FUNCTION_BLOCK PreemptivePriority
VAR_INPUT
  xCondition : ARRAY [1..13] OF BOOL;  (* 条件1 *)
  xTaskComplete : BOOL;  (* 任务完成 *)
  xReset : BOOL;  (* 复位 *)
END_VAR
VAR
  xOccupy : BOOL;  (* 占用 *)
END_VAR
VAR_OUTPUT
  iPriority : INT;  (* 输出任务号 *)
END_VAR
VAR
  m_tonConditionDelay : TON;
  m_xConditionDelay : BOOL;
  m_tConditionCurrentTime : TIME;
  m_iLastTask : INT;  (* 上次执行的任务 *)
  m_tpLastTaskPulse1 : TP;
  m_tpLastTaskPulse2 : TP;
  m_tpLastTaskPulse3 : TP;
  m_tpLastTaskPulse4 : TP;
  m_tpLastTaskPulse5 : TP;
  m_xLastTaskPulse : ARRAY [1..13] OF BOOL;
  m_tLastTaskPulse : ARRAY [1..13] OF TIME := [13(T#0s)];
  m_tpLastTaskPulse6 : TON;
  ii : INT;
END_VAR
VAR CONSTANT
  CONDITION_QUANTITY : INT := 13;
END_VAR
VAR
  m_tpLastTaskPulse7 : TON;
  m_tpLastTaskPulse8 : TON;
  m_tpLastTaskPulse9 : TON;
  m_tpLastTaskPulse10 : TON;
  m_tpLastTaskPulse11 : TON;
  m_tpLastTaskPulse12 : TON;
  m_tpLastTaskPulse13 : TON;
END_VAR
(*抢占式优先级块
现在满足13个条件的任务进行抢占式优先级排列
条件满足后延时两秒，开始执行任务，
同一任务连续执行优先级下降
需要改造成任意多个
使用于一个入口多个出口的程序，使用抢占式优先级块
*)
IF LDP(TRUE, xTaskComplete) THEN
	xOccupy:=0;
	iPriority:=0;
END_IF;
(*//任务滤波，延时两秒*)
m_tonConditionDelay(IN:=( xCondition[1]
						OR xCondition[2]
						OR xCondition[3]
						OR xCondition[4]
						OR xCondition[5]
						OR xCondition[6]
						OR xCondition[7]
						OR xCondition[8]
						OR xCondition[9]
						OR xCondition[10]
						OR xCondition[11]
						OR xCondition[12]
						OR xCondition[13]
						)
						AND iPriority=0,
					PT:= T#1s,
					Q:= m_xConditionDelay ,
					ET:= m_tConditionCurrentTime );		
(*//判断优先级，上个任务与本次任务相同，延时一秒执行*)
m_tpLastTaskPulse1(IN:= xCondition[1]  AND m_iLastTask=1 AND m_xConditionDelay  ,PT:= T#1s,Q:= m_xLastTaskPulse[1],ET:= m_tLastTaskPulse[1] );
m_tpLastTaskPulse2(IN:= xCondition[2]  AND m_iLastTask=2 AND m_xConditionDelay  ,PT:= T#1s,Q:= m_xLastTaskPulse[2],ET:= m_tLastTaskPulse[2] );
m_tpLastTaskPulse3(IN:= xCondition[3]  AND m_iLastTask=3 AND m_xConditionDelay  ,PT:= T#1s,Q:= m_xLastTaskPulse[3],ET:= m_tLastTaskPulse[3] );
m_tpLastTaskPulse4(IN:= xCondition[4]  AND m_iLastTask=4 AND m_xConditionDelay  ,PT:= T#1s,Q:= m_xLastTaskPulse[4],ET:= m_tLastTaskPulse[4] );
m_tpLastTaskPulse5(IN:= xCondition[5]  AND m_iLastTask=5 AND m_xConditionDelay  ,PT:= T#1s,Q:= m_xLastTaskPulse[5],ET:= m_tLastTaskPulse[5] );
m_tpLastTaskPulse6(IN:= xCondition[6]  AND m_iLastTask=6 AND m_xConditionDelay  ,PT:= T#1s,Q:= m_xLastTaskPulse[6],ET:= m_tLastTaskPulse[6] );
m_tpLastTaskPulse7(IN:= xCondition[7]  AND m_iLastTask=7 AND m_xConditionDelay  ,PT:= T#1s,Q:= m_xLastTaskPulse[7],ET:= m_tLastTaskPulse[7] );
m_tpLastTaskPulse8(IN:= xCondition[8]  AND m_iLastTask=8 AND m_xConditionDelay  ,PT:= T#1s,Q:= m_xLastTaskPulse[8],ET:= m_tLastTaskPulse[8] );
m_tpLastTaskPulse9(IN:= xCondition[9]  AND m_iLastTask=9 AND m_xConditionDelay  ,PT:= T#1s,Q:= m_xLastTaskPulse[9],ET:= m_tLastTaskPulse[9] );
m_tpLastTaskPulse10(IN:= xCondition[10]  AND m_iLastTask=10 AND m_xConditionDelay  ,PT:= T#1s,Q:= m_xLastTaskPulse[10],ET:= m_tLastTaskPulse[10] );
m_tpLastTaskPulse11(IN:= xCondition[11]  AND m_iLastTask=11 AND m_xConditionDelay  ,PT:= T#1s,Q:= m_xLastTaskPulse[11],ET:= m_tLastTaskPulse[11] );
m_tpLastTaskPulse12(IN:= xCondition[12]  AND m_iLastTask=12 AND m_xConditionDelay  ,PT:= T#1s,Q:= m_xLastTaskPulse[12],ET:= m_tLastTaskPulse[12] );
m_tpLastTaskPulse13(IN:= xCondition[13]  AND m_iLastTask=13 AND m_xConditionDelay  ,PT:= T#1s,Q:= m_xLastTaskPulse[13],ET:= m_tLastTaskPulse[13] );
(*//执行*)
FOR ii:=1 TO CONDITION_QUANTITY BY 1 DO 
	IF NOT xCondition[ii] AND NOT xOccupy THEN
		iPriority:=0;
	END_IF;
	IF xCondition[ii] AND NOT xOccupy AND m_xConditionDelay AND NOT  m_xLastTaskPulse[ii]  THEN
		iPriority:=ii;
		xOccupy:=1;
		m_iLastTask:=ii;
	END_IF;
END_FOR;        
(*//复位*)
IF xReset THEN
	iPriority:=0;
	xOccupy:=0;
	m_iLastTask:=0;	
END_IF;
(*//清除占用*)
IF iPriority=0 THEN
	xOccupy:=0;
END_IF;
END_FUNCTION_BLOCK

FUNCTION_BLOCK PriorityQueue
VAR_INPUT
  arrxCondition : ARRAY [1..13] OF QueueElement;
  xTaskComplete : BOOL;  (* 任务完成 *)
  xReset : BOOL;  (* 复位 *)
END_VAR
VAR
  xOccupy : BOOL;  (* 占用 *)
END_VAR
VAR_OUTPUT
  iPriority : INT;  (* 输出任务号 *)
END_VAR
VAR
  jj : INT;
END_VAR
VAR CONSTANT
  CONDITION_QUANTITY : INT := 3;
END_VAR
VAR
  arriTaskStack : ARRAY [0..13] OF INT;
  ii : INT;
  kk : INT;
  arrxConditionDelay : ARRAY [1..13] OF BOOL;
  arrxConditionEdgeDetect : ARRAY [1..13] OF BOOL;
  arrxDelayEdgeDetect : ARRAY [1..13] OF BOOL;
  arriDelayCounter : ARRAY [1..13] OF INT;
  ll : INT;
  Temp : INT;
  mm : INT;
  nn : INT;
  Temp2 : INT;
  oo : INT;
END_VAR
(****************************************************************************)
(*
一般情况多对一的任务调度采用这个结构，排队通过出口
优先级功能块，存储任意条件的优先级，实现栈功能先入先出，
复位功能还有问题，
出入栈式优先级块，满足条件后入栈，先入先出，在栈尾加载新任务
栈首为当前执行的任务，任务完成使用上升沿触发，触发后栈首元素弹出

复位功能清空堆栈，栈的容量在CONDITION_QUANTITY 设置
增加了结构体，结构体中带有一个条件函数，和一个优先级指示
任务完成后通过凭借优先级来排序，优先级高的条件先执行   优先级排序是从小到大的，数值小的优先级高
防止干扰，增加了任务的1秒的延时
*)

(***************************************************************************)
(*(//入栈*)
FOR ii:=1 TO CONDITION_QUANTITY BY 1 DO
	(*//循环内无法用定时器，改用计数器的形式*)
	IF arrxCondition[ii].xCondition AND SM411 (*//0.2秒的方波信号，如果移植需要修改成两个定时器*)
		AND arriDelayCounter[ii]<6  (* //计数为6，5个0.2秒的方波，所以为1秒*)
		AND NOT arrxDelayEdgeDetect[ii] THEN    (*//循环内无法用沿函数，增加锁定标志位*)
		arriDelayCounter[ii]:=arriDelayCounter[ii]+1;   (*//计数*)
	END_IF;
	IF NOT arrxCondition[ii].xCondition THEN
		arriDelayCounter[ii]:=0;   (*//计数清零*)
	END_IF;
	arrxDelayEdgeDetect[ii]:=arrxCondition[ii].xCondition AND SM411;  (*//沿函数锁，保证每次SM411为1时只记一次数*)
	IF arriDelayCounter[ii]=5 AND NOT arrxConditionEdgeDetect[ii] THEN;  (*//条件满足1秒后*)
		FOR kk:=0 TO CONDITION_QUANTITY BY 1 DO    
			IF arriTaskStack[kk]=0 THEN
				arriTaskStack[kk]:=ii;   (*//栈尾添加*)
				EXIT;
			END_IF;		
		END_FOR;
	END_IF;	
	arrxConditionEdgeDetect[ii]:=arriDelayCounter[ii]=5;  (*//边沿，这个保证只在=5时，栈尾添加一次*)
END_FOR;
(*//栈顶任务为当前执行的任务**)
iPriority:=arriTaskStack[0]; 
(*//栈顶任务完成，弹出*)
IF 	LDP(TRUE, xTaskComplete) THEN
	FOR jj:=0 TO CONDITION_QUANTITY-1 BY 1 DO
		arriTaskStack[jj]:=arriTaskStack[jj+1];
	END_FOR;
	arriTaskStack[CONDITION_QUANTITY]:=0;(*//栈尾清零*)
	(*//排序，使用插入排序*)
	FOR oo:=0 TO CONDITION_QUANTITY BY 1 DO
		IF arriTaskStack[oo]=0 THEN
			EXIT;  (* //寻找栈中不为零的元素  ，防止0元素进入条件查找的时候报错*)
		END_IF;
	END_FOR;
	(*//插入排序insertionsort*)
	FOR mm:=1 TO oo-1  BY 1 DO   (*//从1开始*)
		Temp:=arriTaskStack[mm];  (*//当前数据记录 *)
		Temp2:=arrxCondition[arriTaskStack[mm]].iPriority;  (*//当前优先级记录 *)
		nn:=mm;  (*//指针赋值*)
		WHILE  (nn>0 AND Temp2< arrxCondition[arriTaskStack[nn-1]].iPriority)  DO  (*//优先级比较，当前优先级小于他前面元素优先级的时候*)
			 arriTaskStack[nn] := arriTaskStack[nn-1] ;  (*//优先级低的向后复制，比TEMP2大的元素都要复制到下一个位置*)
			 nn:=nn-1;
		END_WHILE;
		arriTaskStack[nn]:=Temp; (*//把当前数据放在合适的位置*)
	END_FOR;
END_IF;
(*//复位*)
IF xReset THEN
	FOR jj:=0 TO CONDITION_QUANTITY BY 1 DO
		arriTaskStack[jj]:=0;
	END_FOR;
	FOR ll:=1 TO CONDITION_QUANTITY BY 1 DO
		arrxConditionEdgeDetect[ll]:=0;
		arriDelayCounter[ll]:=0;
	END_FOR;
END_IF;
END_FUNCTION_BLOCK

FUNCTION_BLOCK Conveyor
VAR
  m_xPresentDelay : BOOL;  (* 有无判断延时 *)
  m_xLoadDelayOut : BOOL;  (* 上料延时输出 *)
  m_xInitial : BOOL;  (* 初始化 *)
  m_tUnloadTimer : TIME;  (* 下料计时器 *)
  m_tPresentDelayCurrentTime : TIME;
  m_tonUnloadAlam : TON;  (* 下料报警定时器 *)
  m_tonPresentDelay : TON;  (* 物料有无判断延时，防止误动作 *)
  m_tonNotArriveAlarm : TON;  (* 未到达报警计时 *)
  m_tonLoadDelay : TON;  (* 上料延时 *)
  m_tNotArriveCurrentTime : TIME;  (* 未到达报警计时当前时间 *)
  m_tLoadTimer : TIME;  (* 上料计时器 *)
  iStep : INT;  (* 上料步骤 *)
  m_wStateWord : INT;
END_VAR
VAR_IN_OUT
  ConveyorMotor : ConveyorIO;  (* 输送线输入输出 *)
END_VAR
VAR
  m_tonZoneClear : TON;  (* 初始化清除 *)
  m_tZoneClearCurrentTime : TIME;  (* 初始化清除当前时间 *)
  m_xAutoClear : BOOL;  (* 初始化清除标志位 *)
  m_xZoneClearDone : BOOL;  (* 初始化清除完成 *)
END_VAR
(*////////////////////////////////////////////////////////////////////////////////////////////////////////////
//传输线控制FB块，可控制单方向线体，双向旋转线体，支持双向上下料            
//线体初始化后为空的情况下输入xLoad信号即可进行上料动作，使用xLoadCCW信号可反方向上料
//增加了产品信息和产品种类的储存，当传输线为空和上料进行标志位为零的情况下清除产品信息和产品种类
//使用方式是在置位xLoad信号后，把产品信息和产品种类传入，等下料后自动清零
//线体不为空的情况下使用xUnload信号可进行下料动作，物料有无传感器的下降沿后出发计时器，延时断开传输线旋转
//单方向传输线体把xLoadCCW、xUnloadCCW设置为零，双向线体上料方向和下料反向的,方向固定的 把xUnloadCCW设置为1
//双方向线体双向都能上下料的要根据上料的方向来设置xLoadCCW,xUnloadCCW
//增加工作中信号xBusy当电机正转 显示为工作中
//增加上下料超时报警，xLoadAlarm，xUnloadAlarm，设定时间在LOAD_UNLOAD_TIME常量上，现在设置的为30秒
//增加xPutInto信号，用于直接投入的物料，检测开关感应到后，直接进入下料流程，上升沿有效
//离开延时改为变量 iLeaveDelay 默认为0 离开检测开关离输送线尾端比较远的线体需要根据情况设定100ms为单位
//增加初始化标志位，增加进入延时时间，初始化为进入延时时间为0 ，离开延时时间为2S，通过外围接口可以更改
//修改信息  修改后请增加版本
//12-17进行了优化，增加了未到达报警，当物料未传送到下一设备，就报未到达报警，使用xNextRun标志位制作，没有正常到达
//第0步，不能跳转到第一步把标志位复位，即出现中断情况，2秒后报警
//修改信息  修改后请增加版本
//上料延时增加为50ms防止干扰信号
//nextrun信号在 第三步也要复位
//增加限位报警
//增加超宽报警
//增加产品型号输出在下料的时候把产品型号输送给下一段线体
//增加线体单独复位
//增加任务插入功能配合全局变量
//增加暂停功能
//增加线体状态字显示  0 空闲 1：有料  2 工作中  3  超限报警 4 超宽报警  5 未到达报警  6 下料超时报警
//空料判断放在自动前，进行有无报警判断，然后跳转
//修改超限报警，与尺寸检测报警
////YAO      V1.0
//把所有的IF语句去掉，  IF语句占用指针存储区，容易造成存储区不足的现象
////YAO      V1.1
//初始化清除线体标志位xZoneClear
//ZPA zero pressure accumulation  Term that describes the Conveyor controls and mechanical scheme that will 
//cause loads to queue on a conveyor in discrete zones such that loads do not touch each other(wrapped boxed tray tote carton)
//除了产品信息外，还增加了目标地址，任务类型的数据传递。
//YAO      V1.0
///////////////////////////////////////////////////////////////////////////////////////////////////////////
(*********************************************************)
(*//初始化，
//上料延时位0S，下料报警延时为30S
//下料延时设一个比较大的时间，主要依靠xunload标志位来停止输送线，特殊情况可以用延时来停止物流线下料
//设置时间大的时候计时器会失效*)
IF NOT m_xInitial THEN
	ConveyorMotor.tLoadDelay:=T#100ms;
	ConveyorMotor.tUnloadAlarmDelay:=T#30s;
	ConveyorMotor.xPosLimit:=1;
	ConveyorMotor.xNegLimit:=1;
	ConveyorMotor.xSizeDeficientDetect:=0;
	ConveyorMotor.xZoneClear:=0;
	ConveyorMotor.tZoneClearTime:=T#10s;
	m_xInitial:=1;
END_IF;
(*//自动
//复位信号把步号置0，但xLoad与xUnload没有复位，调用程序需要注意复位后把这两个信号置零，以免发生误动作
//物料有无判断增加延时，防止开自动瞬间误动作发生*)
m_tonPresentDelay(IN:= ConveyorMotor.xCWPresent OR ConveyorMotor.xCCWPresent,
					PT:=T#100ms,
					Q:= m_xPresentDelay,
					ET:= m_tPresentDelayCurrentTime);
CASE iStep OF
0:(*//初始化*)
	ConveyorMotor.xMotorCW:=0;
	ConveyorMotor.xMotorCCW:=0;
	ConveyorMotor.xNextRun:=0;
	ConveyorMotor.iProductCategoryOut:=0;
	ConveyorMotor.iTaskIDOut:=0;
	ConveyorMotor.diDesConveyorOut:=0;
	out(NOT m_xPresentDelay,ConveyorMotor.xEmpty);(*	//判断物料有无传感器*)	
	mov(m_xPresentDelay AND g_xAuto AND NOT ConveyorMotor.xError,3,iStep);(*//自动情况下进行跳转*)(*无超限报警*)
	mov(NOT m_xPresentDelay AND g_xAuto AND NOT ConveyorMotor.xError,1,iStep);
1: (*//上料*)
	rst(ConveyorMotor.xLoad ,ConveyorMotor.iProductCategory);(*//上料开始清除产品信息*)
	rst(ConveyorMotor.xLoad ,ConveyorMotor.iTaskID);
	rst(ConveyorMotor.xLoad ,ConveyorMotor.diDesConveyor);
	mov(ConveyorMotor.xLoad,2,iStep);
2: (*//上料完成*)
	ConveyorMotor.iProductCategory:=ConveyorMotor.iProductCategoryIn;(* //产品信息传入*)
	ConveyorMotor.iTaskID:=ConveyorMotor.iTaskIDIn;
	ConveyorMotor.diDesConveyor:=ConveyorMotor.diDesConveyorIn;
	set(ConveyorMotor.xloadCCW,ConveyorMotor.xMotorCCW);
	rst(ConveyorMotor.xloadCCW,ConveyorMotor.xMotorCW);
	set(NOT ConveyorMotor.xloadCCW,ConveyorMotor.xMotorCW);
	rst(NOT ConveyorMotor.xloadCCW,ConveyorMotor.xMotorCCW);	
	m_tonLoadDelay(IN:= (ConveyorMotor.xCWPresent AND NOT ConveyorMotor.xloadCCW) 
												OR (ConveyorMotor.xCCWPresent AND ConveyorMotor.xloadCCW) ,
										PT:= ConveyorMotor.tLoadDelay ,
										Q:= m_xLoadDelayOut ,
										ET:= m_tLoadTimer );
	mov(m_xLoadDelayOut,3, iStep);
3:(*//下料请求*)	
	ConveyorMotor.xMotorCW:=0;
	ConveyorMotor.xMotorCCW:=0;
	ConveyorMotor.xEmpty:=0;
	mov(ConveyorMotor.xUnload AND NOT ConveyorMotor.xOverWidthAlarm,4,iStep);
4:(*	//下料完成*)
	set(ConveyorMotor.xUnloadCCW,ConveyorMotor.xMotorCCW);
	rst(ConveyorMotor.xUnloadCCW,ConveyorMotor.xMotorCW);
	set(NOT ConveyorMotor.xUnloadCCW,ConveyorMotor.xMotorCW);
	rst(NOT ConveyorMotor.xUnloadCCW,ConveyorMotor.xMotorCCW);	
	ConveyorMotor.xNextRun:=1; (*下一段线体旋转*)
	ConveyorMotor.iProductCategoryOut:=ConveyorMotor.iProductCategory;(*产品型号输出给下一段线体*)
	ConveyorMotor.iTaskIDOut:=ConveyorMotor.iTaskID;
	ConveyorMotor.diDesConveyorOut:=ConveyorMotor.diDesConveyor;
	mov( NOT ConveyorMotor.xUnload , 0, istep );
END_CASE;
(*In-feed zone clear and ready to accept a load from Upstream Conveyor*)
set(ldp(TRUE,g_xAuto) ,m_xAutoClear);
rst(ldf(TRUE,g_xAuto) ,m_xAutoClear);
m_tonZoneClear(IN:= m_xAutoClear AND ConveyorMotor.xZoneClear ,PT:= ConveyorMotor.tZoneClearTime ,Q:=m_xZoneClearDone ,ET:= m_tZoneClearCurrentTime );
set(m_xAutoClear AND ConveyorMotor.xZoneClear,ConveyorMotor.xMotorCW);
mov( m_xAutoClear AND ConveyorMotor.xZoneClear, 0 ,iStep );
rst(  ldf(TRUE, m_xAutoClear ) ,ConveyorMotor.xMotorCW);
rst( m_xZoneClearDone OR m_xPresentDelay  , m_xAutoClear );
(*投入上料，搬出下料，也可用来初始化*)
movp( ConveyorMotor.xPutInto, 0 , iStep );
(*//当前任务显示*)
movp( ConveyorMotor.diDeviceID=g_diDeviceIDSelect , ConveyorMotor.iProductCategory , g_iInsertCategory );
movp( ConveyorMotor.diDeviceID=g_diDeviceIDSelect , ConveyorMotor.iTaskID , g_iInsertTaskID );
dmovp( ConveyorMotor.diDeviceID=g_diDeviceIDSelect , ConveyorMotor.diDesConveyor , g_diInsertDesConveyor );
(*//插入任务*)
mov(g_xInsertTask AND ConveyorMotor.diDeviceID=g_diDeviceIDSelect ,g_iInsertCategory , ConveyorMotor.iProductCategory );
mov(g_xInsertTask AND ConveyorMotor.diDeviceID=g_diDeviceIDSelect , g_iInsertTaskID , ConveyorMotor.iTaskID );
dmov(g_xInsertTask AND ConveyorMotor.diDeviceID=g_diDeviceIDSelect , g_diInsertDesConveyor , ConveyorMotor.diDesConveyor );
(*//单线体复位，当设备号与本线体一致的时候执行复位*)
mov(g_xResetSingle AND ConveyorMotor.diDeviceID=g_diDeviceIDSelect , 0 , iStep );
rst(g_xResetSingle AND ConveyorMotor.diDeviceID=g_diDeviceIDSelect ,ConveyorMotor.xNextRun );
rst(g_xResetSingle AND ConveyorMotor.diDeviceID=g_diDeviceIDSelect  ,ConveyorMotor.xLimitAlarrm );
rst(g_xResetSingle AND ConveyorMotor.diDeviceID=g_diDeviceIDSelect  ,ConveyorMotor.xOverWidthAlarm );
(*//手动*)
(*//正转*)
set( g_xManual 
AND ConveyorMotor.xForward 
AND ConveyorMotor.xBackward=0 
AND ConveyorMotor.xMotorCCW=0 
AND g_xEStop  , 
ConveyorMotor.xMotorCW);
rst((g_xManual 
AND (NOT ConveyorMotor.xForward  
OR ConveyorMotor.xBackward 
OR ConveyorMotor.xMotorCCW )) 
OR NOT g_xEStop,
ConveyorMotor.xMotorCW);
(*//反转*)		
set(g_xManual 
AND ConveyorMotor.xBackward 
AND ConveyorMotor.xForward=0 
AND ConveyorMotor.xMotorCW=0 
AND g_xEStop ,
ConveyorMotor.xMotorCCW);
rst((g_xManual AND 
(NOT ConveyorMotor.xBackward  
OR ConveyorMotor.xForward 
OR ConveyorMotor.xMotorCW ) ) 
OR NOT g_xEStop,
ConveyorMotor.xMotorCCW);
mov(g_xManual ,0,iStep);(*//手动后上下料程序步骤清零*)
(*暂停*)
rst(g_xPause,ConveyorMotor.xMotorCCW);
rst( g_xPause , ConveyorMotor.xMotorCW );
rst(NOT g_xAuto AND NOT g_xManual,ConveyorMotor.xMotorCCW);
rst( NOT g_xAuto AND NOT g_xManual, ConveyorMotor.xMotorCW );
(*工作中信号输出*)
ConveyorMotor.xBusy:=ConveyorMotor.xMotorCCW OR ConveyorMotor.xMotorCW;
(*//未到达报警*)
m_tonNotArriveAlarm(IN:= iStep=0 AND ConveyorMotor.xNextRun  ,PT:= T#2s,Q:= ConveyorMotor.xNotArriveAlarm ,ET:= m_tNotArriveCurrentTime );
(*//下料超时报警*)
m_tonUnloadAlam(IN:= iStep=4,PT:=ConveyorMotor.tUnloadAlarmDelay,Q:= ConveyorMotor.xUnloadAlarm,ET:=m_tUnloadTimer );
(*//限位报警,进料检测开关失效*)
set(  ( ((ConveyorMotor.xloadCCW AND NOT ConveyorMotor.xNegLimit)            (*反转上料，碰到负限位*)
			OR  ( NOT ConveyorMotor.xloadCCW AND NOT ConveyorMotor.xPosLimit)) (*正转上料，碰到正限位*)
		AND iStep=2) (*上料过程*)
	OR
	( iStep=4 (*下料过程*)
		AND( (ConveyorMotor.xUnloadCCW AND NOT ConveyorMotor.xPosLimit)  
			OR (NOT ConveyorMotor.xUnloadCCW AND NOT ConveyorMotor.xNegLimit)))  ,  
	ConveyorMotor.xLimitAlarrm );
mov( ( ((ConveyorMotor.xloadCCW AND NOT ConveyorMotor.xNegLimit)            (*反转上料，碰到负限位*)
			OR  ( NOT ConveyorMotor.xloadCCW AND NOT ConveyorMotor.xPosLimit)) (*正转上料，碰到正限位*)
		AND iStep=2) (*上料过程*)
	OR
	( iStep=4 (*下料过程*)
		AND( (ConveyorMotor.xUnloadCCW AND NOT ConveyorMotor.xPosLimit)  
			OR (NOT ConveyorMotor.xUnloadCCW AND NOT ConveyorMotor.xNegLimit)))  ,
	0,
	iStep);
(*//超宽报警*)
set( (iStep=3 OR iStep=1) AND (NOT ConveyorMotor.xNegLimit OR NOT ConveyorMotor.xPosLimit) , ConveyorMotor.xOverWidthAlarm  );
(*//尺寸不足报警*)
(*//有料状态下检测两个开关都要有信号*)
set( iStep=3 AND ConveyorMotor.xSizeDeficientDetect AND (NOT ConveyorMotor.xCCWPresent OR NOT ConveyorMotor.xCWPresent) ,  ConveyorMotor.xOverWidthAlarm );
mov( iStep=3 AND ConveyorMotor.xSizeDeficientDetect AND (NOT ConveyorMotor.xCCWPresent OR NOT ConveyorMotor.xCWPresent),0,iStep);
(*//总报警*)
ConveyorMotor.xError:=ConveyorMotor.xLimitAlarrm
					OR ConveyorMotor.xNotArriveAlarm
					OR ConveyorMotor.xUnloadAlarm                                             
					OR ConveyorMotor.xOverWidthAlarm;

(*//状态输出*)(*状态显示，容易造成指针容量不足*)
mov( ConveyorMotor.xEmpty AND NOT ConveyorMotor.xBusy , 0 , m_wStateWord);
mov( ConveyorMotor.xEmpty=0 , 							1 , m_wStateWord);
mov( ConveyorMotor.xBusy , 								2 , m_wStateWord);
mov( ConveyorMotor.xLimitAlarrm , 						3, 	m_wStateWord);
mov(ConveyorMotor.xOverWidthAlarm , 					4 , m_wStateWord);
mov( ConveyorMotor.xNotArriveAlarm , 					5 , m_wStateWord);
mov( ConveyorMotor.xUnloadAlarm, 						6 , m_wStateWord);
(*选择本线体后，将状态赋值给全局变量进行显示*)
mov( ConveyorMotor.diDeviceID=g_diDeviceIDSelect , m_wStateWord, g_iConveyorStatus );
END_FUNCTION_BLOCK

PROGRAM TCP
VAR
  m_ton1ReceiveHeartbeat : TON;
  m_t1RecHeartbeatCurrentTime : TIME;
  m_tonAutoClose : TON;
  m_xAutoClose : BOOL;
  m_tAutoCloseCurrentTime : TIME;
  m_tonReconnect : TON;
  m_xReconnect : BOOL;
  m_tReconnectCurrentTime : TIME;
  m_ton5ReceiveHeartbeat : TON;
  m_t5RecHeartbeatCurrentTime : TIME;
  m_ton2ReceiveHeartbeat : TON;
  m_t2RecHeartbeatCurrentTime : TIME;
END_VAR
(*与20通信*)
D200:=2;
(*m_tonReconnect(IN:= NOT SD1282.0 AND NOT SD1284.0,PT:=T#5s  ,Q:=m_xReconnect ,ET:=m_tReconnectCurrentTime);*)
(*1282打开完成状态*)(*1284打开请求状态*)
(*SP_SOCOPEN(m_xReconnect  AND SD1288.A , "U0", K1 , D110 , M100);*)
(*1288.A设备连接状态*)
SP_SOCSND( SM412 AND SD1282.0 , "U0" , K1 , D100, D200, M102 );
SP_SOCRCV( SD1282.0 AND SD1286.0 AND NOT M104 , "U0" , K1, D300 , D400 ,M104 );
(*1286数据接收状态*)
(*m_tonAutoClose(IN:= SD1284.0 AND NOT SD1282.0 ,PT:=T#5s,Q:=m_xAutoClose ,ET:= m_tAutoCloseCurrentTime );
SP_SOCCLOSE( LDF(TRUE,SD1282.0) OR m_xAutoClose  , "U0" , K1, D120, M106 );*)
D201.F:=SM413;
m_ton1ReceiveHeartbeat(IN:=NOT LDP(TRUE, D401.F) ,PT:= t#5S ,Q:= g_x20TcpFailed ,ET:= m_t1RecHeartbeatCurrentTime);
IF g_x20TcpFailed THEN
	M104:=SM413;(*通讯失败有可能是接收模块没动作，重启接收模块*)
	D400:=0;
	D401:=0;
END_IF;



(*与40通信*)
D220:=2;
(*m_tonReconnect(IN:= NOT SD1282.0 AND NOT SD1284.0,PT:=T#5s  ,Q:=m_xReconnect ,ET:=m_tReconnectCurrentTime);*)
(*1282打开完成状态*)(*1284打开请求状态*)
(*SP_SOCOPEN(m_xReconnect  AND SD1288.A , "U0", K1 , D110 , M100);*)
(*1288.A设备连接状态*)
SP_SOCSND( SM412 AND SD1282.4 , "U0" , K5, D120, D220, M122 );
SP_SOCRCV( SD1282.4 AND SD1286.4 AND NOT M124 , "U0" , K5, D320 , D420 ,M124 );
(*1286数据接收状态*)
(*m_tonAutoClose(IN:= SD1284.0 AND NOT SD1282.0 ,PT:=T#5s,Q:=m_xAutoClose ,ET:= m_tAutoCloseCurrentTime );
SP_SOCCLOSE( LDF(TRUE,SD1282.0) OR m_xAutoClose  , "U0" , K1, D120, M106 );*)
D221.F:=SM413;
m_ton2ReceiveHeartbeat(IN:=NOT LDP(TRUE, D421.F) ,PT:= t#5S ,Q:= g_x40TcpFailed ,ET:= m_t2RecHeartbeatCurrentTime);
IF g_x40TcpFailed THEN
	M124:=SM413;(*通讯失败有可能是接收模块没动作，重启接收模块*)
	D420:=0;
	D421:=0;
END_IF;
END_PROGRAM

FUNCTION_BLOCK UConveyor
VAR
  iStep : INT;
END_VAR
VAR_IN_OUT
  ConveyorIOLeft : ConveyorIO;  (* U的左半边 *)
  ConveyorIORight : ConveyorIO;  (* U的右半边 *)
  ConveyorIODown : ConveyorIO;  (* U的下边一横 *)
  UConveyorIO : UConveyorIO;  (* 顶升,阻挡 *)
END_VAR
VAR
  m_xInitial : BOOL;
  m_tonCylinderOvertime : TON;  (* 气缸超时报警定时器 *)
  m_tCylinderOvertimeCurrent : TIME;
  m_tonExitBarDelay : TON;  (* 退出阻挡器延时 *)
  m_tExitBarDelay : TIME;
  m_xExitBarDelay : BOOL;
END_VAR
(*                                                                                                          
初始化中增加气缸复位，气缸位置有BUG
//*)
IF NOT m_xInitial THEN
		UConveyorIO.tSetOvertime:=T#5s;
	UConveyorIO.xExitEnable1:=1;
	UConveyorIO.xExitEnable2:=1;
	UConveyorIO.xExitEnable3:=1;
	m_xInitial:=1;
END_IF;
(*外部不用写ConveyorDown的开关，会自己根据来料的产品信息判断停哪个光电*)
IF UConveyorIO.iTask=1 AND ConveyorIODown.diDesConveyorIn=ConveyorIOLeft.diDeviceID THEN
	ConveyorIODown.xCWPresent:=ConveyorIOLeft.xCCWPresent;
ELSIF UConveyorIO.iTask=1 AND ConveyorIODown.diDesConveyorIn=ConveyorIORight.diDeviceID THEN
	ConveyorIODown.xCWPresent:=ConveyorIORight.xCCWPresent;
ELSE
	ConveyorIODown.xCWPresent:=ConveyorIOLeft.xCCWPresent OR ConveyorIORight.xCCWPresent;
END_IF;
(*这里判断什么时候直接放行，左右都不需要，也不是0，就放走*)
IF  NOT(ConveyorIODown.diDesConveyor=ConveyorIOLeft.diDeviceID 
		OR  ConveyorIODown.diDesConveyor=ConveyorIORight.diDeviceID 
		OR ConveyorIODown.diDesConveyor=0) THEN
	UConveyorIO.xPassEnable:=1;
ELSE
	UConveyorIO.xPassEnable:=0;
END_IF;	
IF g_xAuto THEN	
(*	//加个Step为0的延时，防止扫描周期的影响*)
	m_TonStep0(IN:= iStep=0 ,PT:= t#100ms ,Q:= m_xStep0 ,ET:= m_tStep0 );
	(*//这个是留给阻挡动作的时间*)
	m_tonExitBarDelay(IN:=iStep=4 ,PT:= T#1s ,Q:= m_xExitBarDelay ,ET:= m_tExitBarDelay);
CASE UConveyorIO.iTask OF(*这个Task做抢占，可做LastTask保护*)
0:(*各种初始化，能自动去3*)
	ConveyorIODown.xLoad:=0;
	ConveyorIOleft.xLoad:=0;
	ConveyorIORight.xLoad:=0;
	ConveyorIODown.xUnload:=0;
	ConveyorIOLeft.xUnload:=0;
	ConveyorIORight.xUnload:=0;
	ConveyorIODown.xPutInto:=0;
	ConveyorIOLeft.xPutInto:=0;
	ConveyorIORight.xPutInto:=0;	
	UConveyorIO.xExitBarCylinderRetract1:=0;
	UConveyorIO.xExitBarCylinderRetract2:=0;	
	UConveyorIO.xLiftCylinderRetract1:=1;
	UConveyorIO.xLiftCylinderRetract2:=1;
	UConveyorIO.xLiftCylinderExtend1:=0;
	UConveyorIO.xLiftCylinderExtend2:=0;
1:(*上料*)
	CASE iStep OF
	0:(*各种初始化，能自动去3*)
		ConveyorIODown.xLoad:=0;
		ConveyorIOleft.xLoad:=0;
		ConveyorIORight.xLoad:=0;
		ConveyorIODown.xUnload:=0;
		ConveyorIOLeft.xUnload:=0;
		ConveyorIORight.xUnload:=0;
		UConveyorIO.xExitBarCylinderRetract1:=0;
		UConveyorIO.xExitBarCylinderRetract2:=0;
		UConveyorIO.xBatteryError:=0;
		ConveyorIODown.xPutInto:=0;
		ConveyorIOLeft.xPutInto:=0;
		ConveyorIORight.xPutInto:=0;	
	(*	//根据是否有料判断去1还是3，但会等一个延时*)
		IF m_xStep0 AND  ConveyorIODown.xEmpty THEN
			iStep:=1;
		ELSIF m_xStep0 AND NOT ConveyorIODown.xEmpty THEN
			iStep:=3;
		END_IF;	
	1:(*顶升初始化，等load*)
		(*//左顶升*)
		IF UConveyorIO.xLiftCylinderExtendInit1 THEN
			UConveyorIO.xLiftCylinderExtend1:=1;
			UConveyorIO.xLiftCylinderRetract1:=0;
		ELSE
			UConveyorIO.xLiftCylinderExtend1:=0;
			UConveyorIO.xLiftCylinderRetract1:=1;
		END_IF;
	(*	//右顶升*)
		IF UConveyorIO.xLiftCylinderExtendInit2 THEN
			UConveyorIO.xLiftCylinderExtend2:=1;
			UConveyorIO.xLiftCylinderRetract2:=0;
			ELSE
			UConveyorIO.xLiftCylinderExtend2:=0;
			UConveyorIO.xLiftCylinderRetract2:=1;
		END_IF;
		(*//顶升到位，等上料信号*)
		IF 	((UConveyorIO.xLiftCylinderExtendInit1 AND UConveyorIO.xLiftCylinderExtendDetect1)
				OR (NOT UConveyorIO.xLiftCylinderExtendInit1 AND UConveyorIO.xLiftCylinderRetractDetect1))
			AND	((UConveyorIO.xLiftCylinderExtendInit2 AND UConveyorIO.xLiftCylinderExtendDetect2)
		   		OR (NOT UConveyorIO.xLiftCylinderExtendInit2 AND UConveyorIO.xLiftCylinderRetractDetect2))		
			AND	UConveyorIO.xEntryEnable1 THEN(*有上料请求1*)
		   	ConveyorIODown.xLoad:=1;
			iStep:=2;
		END_IF;
	2:(*Load完成*)
		(*去右臂时才需要阻挡1放行,其他情况阻挡1挡住*)
		UConveyorIO.xExitBarCylinderRetract1:=ConveyorIODown.diDesConveyorIn=ConveyorIORight.diDeviceID;
		IF NOT ConveyorIODown.xEmpty THEN
			ConveyorIODown.xLoad:=0;
			ConveyorIOLeft.xPutInto:=1;
			ConveyorIOright.xPutInto:=1;
			istep:=3;
		END_IF;
	3:(*顶升等Unload，这里等有了ExitEnable再顶升，因为可能有地方需要允许了再升降，比如倍速链*)
		(*//电池检测保护，防止把带电池的料框送进去了*)
		IF (ConveyorIODown.diDesConveyor=ConveyorIOLeft.diDeviceID OR ConveyorIODown.diDesConveyor=ConveyorIORight.diDeviceID)
			AND	(UConveyorIO.xBatteryDetect1 OR UConveyorIO.xBatteryDetect2)(*在下面时检测*)
			AND UConveyorIO.xLiftCylinderRetractDetect1 AND UConveyorIO.xLiftCylinderRetractDetect2 THEN
			UConveyorIO.xBatteryError:=1;
		END_IF;	
		(*//左侧顶升控制*)
		IF (ConveyorIODown.diDesConveyor=ConveyorIOLeft.diDeviceID AND UConveyorIO.xExitEnable2 AND NOT UConveyorIO.xBatteryError)THEN
			IF UConveyorIO.xLiftCylinderExtendInit1 THEN
				UConveyorIO.xLiftCylinderExtend1:=0;
				UConveyorIO.xLiftCylinderRetract1:=1;
			ELSE
				UConveyorIO.xLiftCylinderExtend1:=1;
				UConveyorIO.xLiftCylinderRetract1:=0;
			END_IF;
			IF(NOT UConveyorIO.xLiftCylinderExtendInit1 AND UConveyorIO.xLiftCylinderExtendDetect1)
				OR (UConveyorIO.xLiftCylinderExtendInit1 AND UConveyorIO.xLiftCylinderRetractDetect1)THEN
				ConveyorIOLeft.xPutInto:=0;
				ConveyorIOright.xPutInto:=0;
				iStep:=4;
			END_IF;
		END_IF;	
		(*//右侧顶升控制*)
		IF (ConveyorIODown.diDesConveyor=ConveyorIORight.diDeviceID AND UConveyorIO.xExitEnable3 AND NOT UConveyorIO.xBatteryError)THEN
			IF UConveyorIO.xLiftCylinderExtendInit2 THEN
				UConveyorIO.xLiftCylinderExtend2:=0;
				UConveyorIO.xLiftCylinderRetract2:=1;
			ELSE
				UConveyorIO.xLiftCylinderExtend2:=1;
				UConveyorIO.xLiftCylinderRetract2:=0;
			END_IF;
			IF(NOT UConveyorIO.xLiftCylinderExtendInit2 AND UConveyorIO.xLiftCylinderExtendDetect2)
				OR (UConveyorIO.xLiftCylinderExtendInit2 AND UConveyorIO.xLiftCylinderRetractDetect2) THEN
				ConveyorIOLeft.xPutInto:=0;
				ConveyorIOright.xPutInto:=0;
				iStep:=4;
			END_IF;
		END_IF;	
	(*	//直接放行控制*)
		IF UConveyorIO.xPassEnable AND UConveyorIO.xExitEnable1 AND NOT UConveyorIO.xBatteryError THEN
			IF UConveyorIO.xLiftCylinderExtendInit1 THEN
				UConveyorIO.xLiftCylinderExtend1:=1;
				UConveyorIO.xLiftCylinderRetract1:=0;
			ELSE
				UConveyorIO.xLiftCylinderExtend1:=0;
				UConveyorIO.xLiftCylinderRetract1:=1;
			END_IF;
			IF UConveyorIO.xLiftCylinderExtendInit2 THEN
				UConveyorIO.xLiftCylinderExtend2:=1;
				UConveyorIO.xLiftCylinderRetract2:=0;
			ELSE
				UConveyorIO.xLiftCylinderExtend2:=0;
				UConveyorIO.xLiftCylinderRetract2:=1;
			END_IF;
			IF((UConveyorIO.xLiftCylinderExtendInit1 AND UConveyorIO.xLiftCylinderExtendDetect1)
 OR (NOT UConveyorIO.xLiftCylinderExtendInit1 AND UConveyorIO.xLiftCylinderRetractDetect1))
				AND((UConveyorIO.xLiftCylinderExtendInit2 AND UConveyorIO.xLiftCylinderExtendDetect2)
 OR (NOT UConveyorIO.xLiftCylinderExtendInit2 AND UConveyorIO.xLiftCylinderRetractDetect2))THEN
				UConveyorIO.xExitBarCylinderRetract1:=1;
				UConveyorIO.xExitBarCylinderRetract2:=1;
				ConveyorIOLeft.xPutInto:=0;
				ConveyorIOright.xPutInto:=0;
				iStep:=4;
			END_IF;	
		END_IF;
	4:(*Unload完成，回0*)
			IF ConveyorIODown.diDesConveyor=ConveyorIOLeft.diDeviceID AND UConveyorIO.xExitEnable2 AND m_xExitBarDelay THEN
				ConveyorIOLeft.xUnload:=1;
			ELSIF ConveyorIODown.diDesConveyor=ConveyorIORight.diDeviceID AND UConveyorIO.xExitEnable3 AND m_xExitBarDelay THEN
				ConveyorIORight.xUnload:=1;
			ELSIF UConveyorIO.xPassEnable AND UConveyorIO.xExitEnable1 AND m_xExitBarDelay THEN
				ConveyorIODown.xUnload:=1;
			ELSE
				ConveyorIODown.xUnload:=0;
				ConveyorIOLeft.xUnload:=0;
				ConveyorIORight.xUnload:=0;
			END_IF;	
		IF ( (ConveyorIODown.diDesConveyor=ConveyorIOLeft.diDeviceID  AND LDF(TRUE,UConveyorIO.xExitEnable2))
		  OR(ConveyorIODown.diDesConveyor=ConveyorIORight.diDeviceID AND LDF(TRUE,UConveyorIO.xExitEnable3))
		  OR(UConveyorIO.xPassEnable AND LDF(TRUE,UConveyorIO.xExitEnable1)) )AND m_xExitBarDelay  THEN
			ConveyorIODown.xUnload:=0;
			ConveyorIOLeft.xUnload:=0;
			ConveyorIORight.xUnload:=0;
			ConveyorIODown.xPutInto:=1;
			ConveyorIOLeft.xPutInto:=1;
			ConveyorIORight.xPutInto:=1;
			UConveyorIO.xExitBarCylinderRetract1:=0;
			UConveyorIO.xExitBarCylinderRetract2:=0;
			iStep:=0;
		END_IF;
	END_CASE;
2:(*左下料*)
	CASE iStep OF
	0:(*各种初始化，能自动去3*)
		ConveyorIODown.xLoad:=0;
		ConveyorIOleft.xLoad:=0;
		ConveyorIORight.xLoad:=0;
		ConveyorIODown.xUnload:=0;
		ConveyorIOLeft.xUnload:=0;
		ConveyorIORight.xUnload:=0;
		UConveyorIO.xBatteryError:=0;
		UConveyorIO.xExitBarCylinderRetract1:=0;
		UConveyorIO.xExitBarCylinderRetract2:=0;
		ConveyorIODown.xPutInto:=0;
		ConveyorIOLeft.xPutInto:=0;
		ConveyorIORight.xPutInto:=0;
		IF m_xStep0 AND  ConveyorIODown.xEmpty THEN
			iStep:=1;
		ELSIF m_xStep0 AND NOT ConveyorIODown.xEmpty THEN
			iStep:=3;
		END_IF;	
	1:(*左顶升动作，等load*)
		IF UConveyorIO.xLiftCylinderExtendInit1 THEN
			UConveyorIO.xLiftCylinderExtend1:=0;
			UConveyorIO.xLiftCylinderRetract1:=1;
			ELSE
			UConveyorIO.xLiftCylinderExtend1:=1;
			UConveyorIO.xLiftCylinderRetract1:=0;
		END_IF;
		IF ((NOT UConveyorIO.xLiftCylinderExtendInit1 AND UConveyorIO.xLiftCylinderExtendDetect1)
			OR ( UConveyorIO.xLiftCylinderExtendInit1 AND UConveyorIO.xLiftCylinderRetractDetect1))
			AND UConveyorIO.xEntryEnable2 THEN(*有上料请求1*)
		   	ConveyorIOLeft.xLoad:=1;
			iStep:=2;
		END_IF;
	2:(*Load完成*)
		IF NOT ConveyorIOLeft.xEmpty THEN
			ConveyorIOLeft.xLoad:=0;
			ConveyorIODown.xPutInto:=1;
			ConveyorIODown.diDesConveyor:=ConveyorIOLeft.diDesConveyor;
			istep:=3;
		END_IF;
	3:(*顶升等Unload，这里等有了ExitEnable再顶升，因为可能有地方需要允许了再升降，比如倍速链*)
		UConveyorIO.xExitBarCylinderRetract1:=1;
		UConveyorIO.xExitBarCylinderRetract2:=1;
		IF  UConveyorIO.xExitEnable1 THEN
			IF UConveyorIO.xLiftCylinderExtendInit1 THEN
				UConveyorIO.xLiftCylinderExtend1:=1;
				UConveyorIO.xLiftCylinderRetract1:=0;
			ELSE
				UConveyorIO.xLiftCylinderExtend1:=0;
				UConveyorIO.xLiftCylinderRetract1:=1;
			END_IF;
			IF(( UConveyorIO.xLiftCylinderExtendInit1 AND UConveyorIO.xLiftCylinderExtendDetect1)